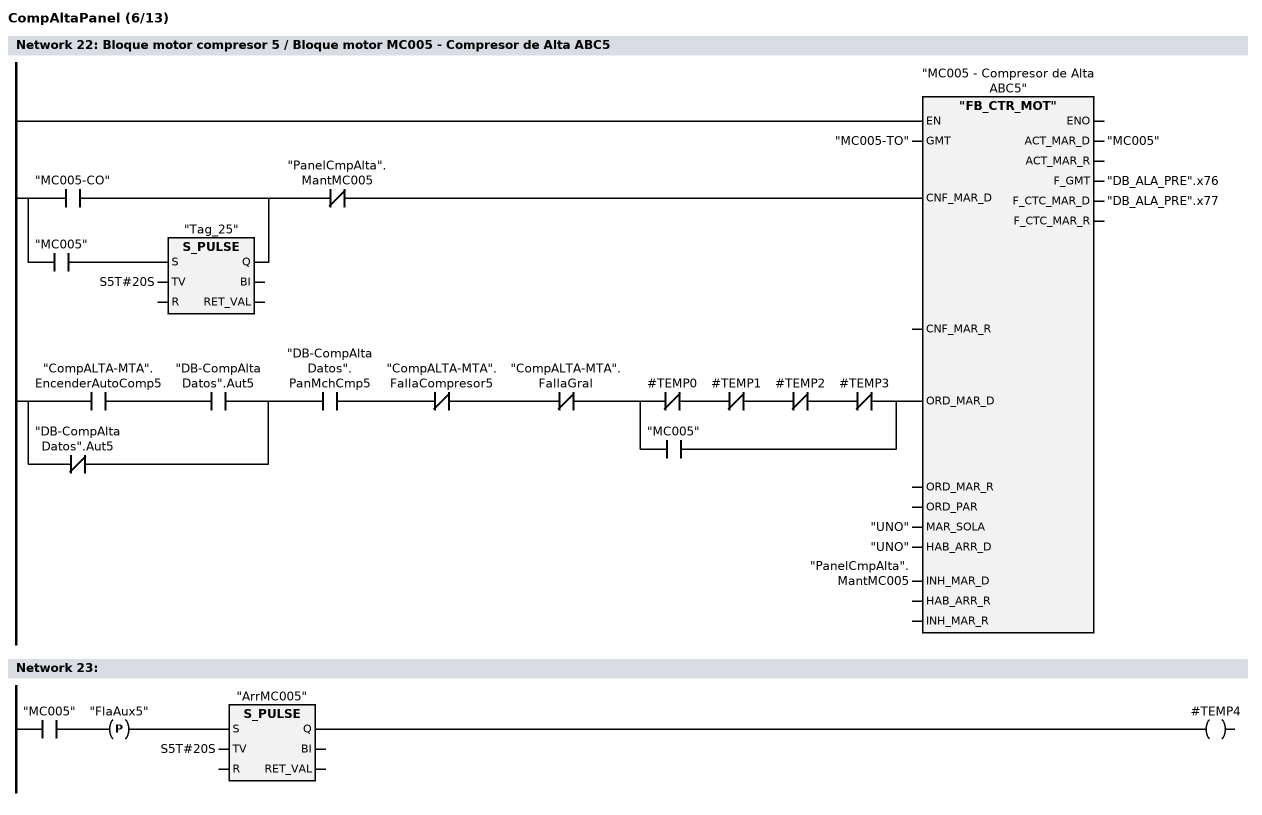
   RUNG wire#powerrail
      "MC005 - Compresor de Alta ABC5"(CNF_MAR_D := wire#w2, ORD_MAR_D := wire#w5, GMT := "MC005-TO", CNF_MAR_R :=, ORD_MAR_R :=, ORD_PAR :=, MAR_SOLA := "UNO", HAB_ARR_D := "UNO", INH_MAR_D := "PanelCmpAlta".MantMC005, HAB_ARR_R :=, INH_MAR_R :=, ACT_MAR_D => "MC005", ACT_MAR_R =>, F_GMT => "DB_ALA_PRE".x76, F_CTC_MAR_D => "DB_ALA_PRE".x77, F_CTC_MAR_R =>)
   END_RUNG
   RUNG wire#powerrail
      Contact( "MC005-CO" )
      wire#w1
      I_Contact( "PanelCmpAlta".MantMC005 )
   END_RUNG wire#w2
   RUNG wire#powerrail
      Contact( "MC005" )
      S_PULSE(T_NO := "Tag_25", TV := S5T#20S, R :=, BI =>, RET_VAL =>)
   END_RUNG wire#w1
   RUNG wire#powerrail
      Contact( "CompALTA-MTA".EncenderAutoComp5 )
      Contact( "DB-CompAltaDatos".Aut5 )
      wire#w3
      Contact( "DB-CompAltaDatos".PanMchCmp5 )
      I_Contact( "CompALTA-MTA".FallaCompresor5 )
      I_Contact( "CompALTA-MTA".FallaGral )
      wire#w4
      I_Contact( #TEMP0 )
      I_Contact( #TEMP1 )
      I_Contact( #TEMP2 )
      I_Contact( #TEMP3 )
   END_RUNG wire#w5
   RUNG wire#powerrail
      I_Contact( "DB-CompAltaDatos".Aut5 )
   END_RUNG wire#w3
   RUNG wire#w4
      Contact( "MC005" )
   END_RUNG wire#w5
   // the same network as SCL:
   #_s5time1 := S_PULSE(T_NO := "Tag_25", S := "MC005", TV := S5T#20S, Q => #_w1);
   "MC005 - Compresor de Alta ABC5"(GMT := "MC005-TO",   // "FB_CTR_MOT"
                           CNF_MAR_D := ("MC005-CO" OR #_w1) AND NOT "PanelCmpAlta".MantMC005,
                           ORD_MAR_D := (("CompALTA-MTA".EncenderAutoComp5 AND "DB-CompAltaDatos".Aut5) OR NOT "DB-CompAltaDatos".Aut5) AND "DB-CompAltaDatos".PanMchCmp5 AND NOT "CompALTA-MTA".FallaCompresor5 AND NOT "CompALTA-MTA".FallaGral AND ((NOT #TEMP0 AND NOT #TEMP1 AND NOT #TEMP2 AND NOT #TEMP3) OR "MC005"),
                           MAR_SOLA := "UNO",
                           HAB_ARR_D := "UNO",
                           INH_MAR_D := "PanelCmpAlta".MantMC005,
                           ACT_MAR_D => "MC005",
                           F_GMT => "DB_ALA_PRE".x76,
                           F_CTC_MAR_D => "DB_ALA_PRE".x77);
END_REGION

REGION Network 23
   RUNG wire#powerrail
      Contact( "MC005" )
      P_Trig( "FlaAux5" )
      S_PULSE(T_NO := "ArrMC005", TV := S5T#20S, R :=, BI =>, RET_VAL =>)
      Coil( #TEMP4 )
   END_RUNG
   // the same network as SCL:
   #_w1 := "MC005" AND NOT "FlaAux5";   // rising edge
   "FlaAux5" := "MC005";
   #_s5time1 := S_PULSE(T_NO := "ArrMC005", S := #_w1, TV := S5T#20S, Q => #_w2);
   #TEMP4 := #_w2;
END_REGION

REGION Network 24: Bloque motor compresor 6 / Bloque motor MC005 - Compresor de Alta ABC5
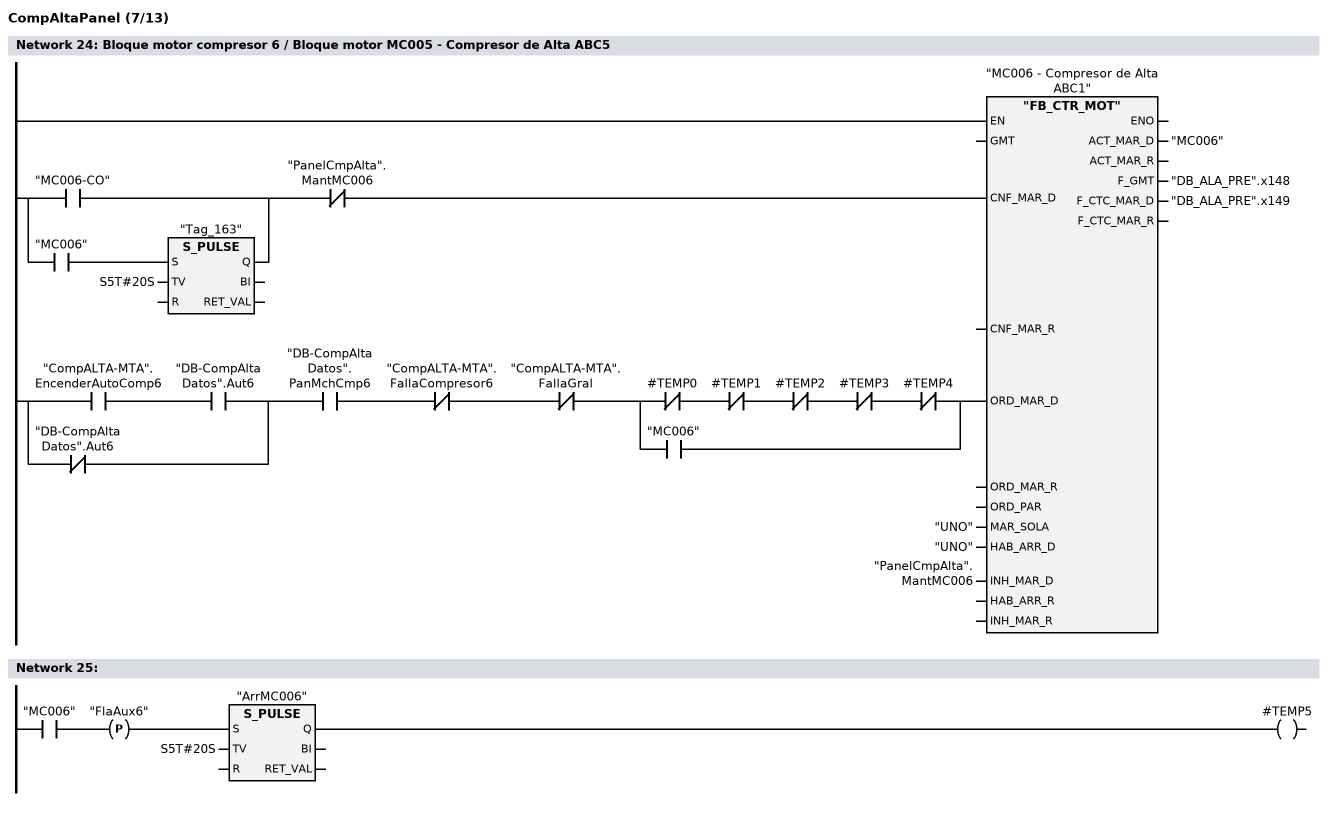
   RUNG wire#powerrail
      "MC006 - Compresor de Alta ABC1"(CNF_MAR_D := wire#w2, ORD_MAR_D := wire#w5, GMT :=, CNF_MAR_R :=, ORD_MAR_R :=, ORD_PAR :=, MAR_SOLA := "UNO", HAB_ARR_D := "UNO", INH_MAR_D := "PanelCmpAlta".MantMC006, HAB_ARR_R :=, INH_MAR_R :=, ACT_MAR_D => "MC006", ACT_MAR_R =>, F_GMT => "DB_ALA_PRE".x148, F_CTC_MAR_D => "DB_ALA_PRE".x149, F_CTC_MAR_R =>)
   END_RUNG
   RUNG wire#powerrail
      Contact( "MC006-CO" )
      wire#w1
      I_Contact( "PanelCmpAlta".MantMC006 )
   END_RUNG wire#w2
   RUNG wire#powerrail
      Contact( "MC006" )
      S_PULSE(T_NO := "Tag_163", TV := S5T#20S, R :=, BI =>, RET_VAL =>)
   END_RUNG wire#w1
   RUNG wire#powerrail
      Contact( "CompALTA-MTA".EncenderAutoComp6 )
      Contact( "DB-CompAltaDatos".Aut6 )
      wire#w3
      Contact( "DB-CompAltaDatos".PanMchCmp6 )
      I_Contact( "CompALTA-MTA".FallaCompresor6 )
      I_Contact( "CompALTA-MTA".FallaGral )
      wire#w4
      I_Contact( #TEMP0 )
      I_Contact( #TEMP1 )
      I_Contact( #TEMP2 )
      I_Contact( #TEMP3 )
      I_Contact( #TEMP4 )
   END_RUNG wire#w5
   RUNG wire#powerrail
      I_Contact( "DB-CompAltaDatos".Aut6 )
   END_RUNG wire#w3
   RUNG wire#w4
      Contact( "MC006" )
   END_RUNG wire#w5
   // the same network as SCL:
   #_s5time1 := S_PULSE(T_NO := "Tag_163", S := "MC006", TV := S5T#20S, Q => #_w1);
   "MC006 - Compresor de Alta ABC1"(CNF_MAR_D := ("MC006-CO" OR #_w1) AND NOT "PanelCmpAlta".MantMC006,   // "FB_CTR_MOT"
                           ORD_MAR_D := (("CompALTA-MTA".EncenderAutoComp6 AND "DB-CompAltaDatos".Aut6) OR NOT "DB-CompAltaDatos".Aut6) AND "DB-CompAltaDatos".PanMchCmp6 AND NOT "CompALTA-MTA".FallaCompresor6 AND NOT "CompALTA-MTA".FallaGral AND ((NOT #TEMP0 AND NOT #TEMP1 AND NOT #TEMP2 AND NOT #TEMP3 AND NOT #TEMP4) OR "MC006"),
                           MAR_SOLA := "UNO",
                           HAB_ARR_D := "UNO",
                           INH_MAR_D := "PanelCmpAlta".MantMC006,
                           ACT_MAR_D => "MC006",
                           F_GMT => "DB_ALA_PRE".x148,
                           F_CTC_MAR_D => "DB_ALA_PRE".x149);
END_REGION

REGION Network 25
   RUNG wire#powerrail
      Contact( "MC006" )
      P_Trig( "FlaAux6" )
      S_PULSE(T_NO := "ArrMC006", TV := S5T#20S, R :=, BI =>, RET_VAL =>)
      Coil( #TEMP5 )
   END_RUNG
   // the same network as SCL:
   #_w1 := "MC006" AND NOT "FlaAux6";   // rising edge
   "FlaAux6" := "MC006";
   #_s5time1 := S_PULSE(T_NO := "ArrMC006", S := #_w1, TV := S5T#20S, Q => #_w2);
   #TEMP5 := #_w2;
END_REGION

REGION Network 26: Bloque de animación motor compresor 1 / Animación Motor MC001 - Compresor de Alta ABC2
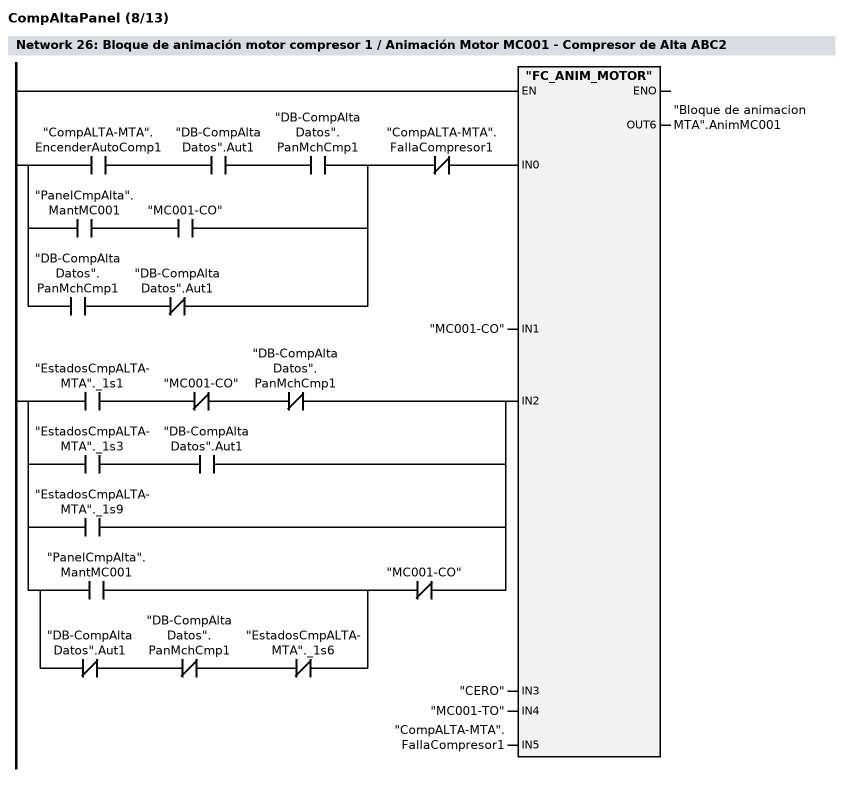
   RUNG wire#powerrail
      "FC_ANIM_MOTOR"(IN0 := wire#w2, IN2 := wire#w4, IN1 := "MC001-CO", IN3 := "CERO", IN4 := "MC001-TO", IN5 := "CompALTA-MTA".FallaCompresor1, OUT6 => "Bloque de animacion MTA".AnimMC001)
   END_RUNG
   RUNG wire#powerrail
      Contact( "CompALTA-MTA".EncenderAutoComp1 )
      Contact( "DB-CompAltaDatos".Aut1 )
      Contact( "DB-CompAltaDatos".PanMchCmp1 )
      wire#w1
      I_Contact( "CompALTA-MTA".FallaCompresor1 )
   END_RUNG wire#w2
   RUNG wire#powerrail
      Contact( "PanelCmpAlta".MantMC001 )
      Contact( "MC001-CO" )
   END_RUNG wire#w1
   RUNG wire#powerrail
      Contact( "DB-CompAltaDatos".PanMchCmp1 )
      I_Contact( "DB-CompAltaDatos".Aut1 )
   END_RUNG wire#w1
   RUNG wire#powerrail
      Contact( "EstadosCmpALTA-MTA"._1s1 )
      I_Contact( "MC001-CO" )
      I_Contact( "DB-CompAltaDatos".PanMchCmp1 )
   END_RUNG wire#w4
   RUNG wire#powerrail
      Contact( "EstadosCmpALTA-MTA"._1s3 )
      Contact( "DB-CompAltaDatos".Aut1 )
   END_RUNG wire#w4
   RUNG wire#powerrail
      Contact( "EstadosCmpALTA-MTA"._1s9 )
   END_RUNG wire#w4
   RUNG wire#powerrail
      Contact( "PanelCmpAlta".MantMC001 )
      wire#w3
      I_Contact( "MC001-CO" )
   END_RUNG wire#w4
   RUNG wire#powerrail
      I_Contact( "DB-CompAltaDatos".Aut1 )
      I_Contact( "DB-CompAltaDatos".PanMchCmp1 )
      I_Contact( "EstadosCmpALTA-MTA"._1s6 )
   END_RUNG wire#w3
   // the same network as SCL:
   "FC_ANIM_MOTOR"(IN0 := (("CompALTA-MTA".EncenderAutoComp1 AND "DB-CompAltaDatos".Aut1 AND "DB-CompAltaDatos".PanMchCmp1) OR ("PanelCmpAlta".MantMC001 AND "MC001-CO") OR ("DB-CompAltaDatos".PanMchCmp1 AND NOT "DB-CompAltaDatos".Aut1)) AND NOT "CompALTA-MTA".FallaCompresor1,
                   IN1 := "MC001-CO",
                   IN2 := ("EstadosCmpALTA-MTA"._1s1 AND NOT "MC001-CO" AND NOT "DB-CompAltaDatos".PanMchCmp1) OR ("EstadosCmpALTA-MTA"._1s3 AND "DB-CompAltaDatos".Aut1) OR "EstadosCmpALTA-MTA"._1s9 OR (("PanelCmpAlta".MantMC001 OR (NOT "DB-CompAltaDatos".Aut1 AND NOT "DB-CompAltaDatos".PanMchCmp1 AND NOT "EstadosCmpALTA-MTA"._1s6)) AND NOT "MC001-CO"),
                   IN3 := "CERO",
                   IN4 := "MC001-TO",
                   IN5 := "CompALTA-MTA".FallaCompresor1,
                   OUT6 => "Bloque de animacion MTA".AnimMC001);
END_REGION

REGION Network 27: Bloque de animación motor compresor 2 / Animación Motor MC002 - Compresor de Alta ABC3
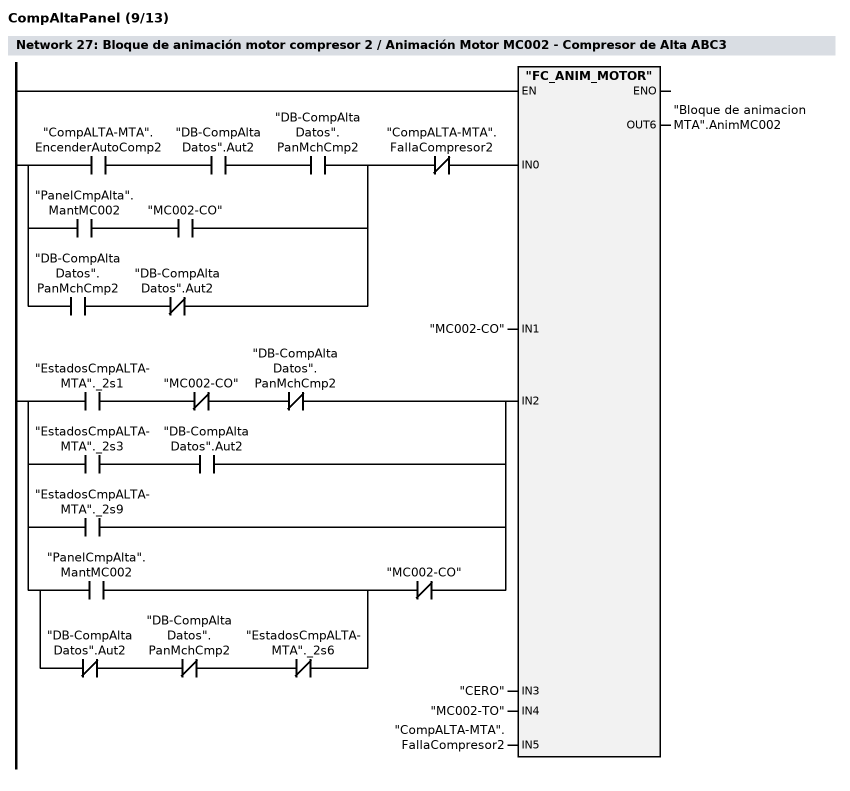
   RUNG wire#powerrail
      "FC_ANIM_MOTOR"(IN0 := wire#w2, IN2 := wire#w4, IN1 := "MC002-CO", IN3 := "CERO", IN4 := "MC002-TO", IN5 := "CompALTA-MTA".FallaCompresor2, OUT6 => "Bloque de animacion MTA".AnimMC002)
   END_RUNG
   RUNG wire#powerrail
      Contact( "CompALTA-MTA".EncenderAutoComp2 )
      Contact( "DB-CompAltaDatos".Aut2 )
      Contact( "DB-CompAltaDatos".PanMchCmp2 )
      wire#w1
      I_Contact( "CompALTA-MTA".FallaCompresor2 )
   END_RUNG wire#w2
   RUNG wire#powerrail
      Contact( "PanelCmpAlta".MantMC002 )
      Contact( "MC002-CO" )
   END_RUNG wire#w1
   RUNG wire#powerrail
      Contact( "DB-CompAltaDatos".PanMchCmp2 )
      I_Contact( "DB-CompAltaDatos".Aut2 )
   END_RUNG wire#w1
   RUNG wire#powerrail
      Contact( "EstadosCmpALTA-MTA"._2s1 )
      I_Contact( "MC002-CO" )
      I_Contact( "DB-CompAltaDatos".PanMchCmp2 )
   END_RUNG wire#w4
   RUNG wire#powerrail
      Contact( "EstadosCmpALTA-MTA"._2s3 )
      Contact( "DB-CompAltaDatos".Aut2 )
   END_RUNG wire#w4
   RUNG wire#powerrail
      Contact( "EstadosCmpALTA-MTA"._2s9 )
   END_RUNG wire#w4
   RUNG wire#powerrail
      Contact( "PanelCmpAlta".MantMC002 )
      wire#w3
      I_Contact( "MC002-CO" )
   END_RUNG wire#w4
   RUNG wire#powerrail
      I_Contact( "DB-CompAltaDatos".Aut2 )
      I_Contact( "DB-CompAltaDatos".PanMchCmp2 )
      I_Contact( "EstadosCmpALTA-MTA"._2s6 )
   END_RUNG wire#w3
   // the same network as SCL:
   "FC_ANIM_MOTOR"(IN0 := (("CompALTA-MTA".EncenderAutoComp2 AND "DB-CompAltaDatos".Aut2 AND "DB-CompAltaDatos".PanMchCmp2) OR ("PanelCmpAlta".MantMC002 AND "MC002-CO") OR ("DB-CompAltaDatos".PanMchCmp2 AND NOT "DB-CompAltaDatos".Aut2)) AND NOT "CompALTA-MTA".FallaCompresor2,
                   IN1 := "MC002-CO",
                   IN2 := ("EstadosCmpALTA-MTA"._2s1 AND NOT "MC002-CO" AND NOT "DB-CompAltaDatos".PanMchCmp2) OR ("EstadosCmpALTA-MTA"._2s3 AND "DB-CompAltaDatos".Aut2) OR "EstadosCmpALTA-MTA"._2s9 OR (("PanelCmpAlta".MantMC002 OR (NOT "DB-CompAltaDatos".Aut2 AND NOT "DB-CompAltaDatos".PanMchCmp2 AND NOT "EstadosCmpALTA-MTA"._2s6)) AND NOT "MC002-CO"),
                   IN3 := "CERO",
                   IN4 := "MC002-TO",
                   IN5 := "CompALTA-MTA".FallaCompresor2,
                   OUT6 => "Bloque de animacion MTA".AnimMC002);
END_REGION

REGION Network 28: Bloque de animación motor compresor 3 / Animación Motor MC003 - Compresor de Alta BELLIS
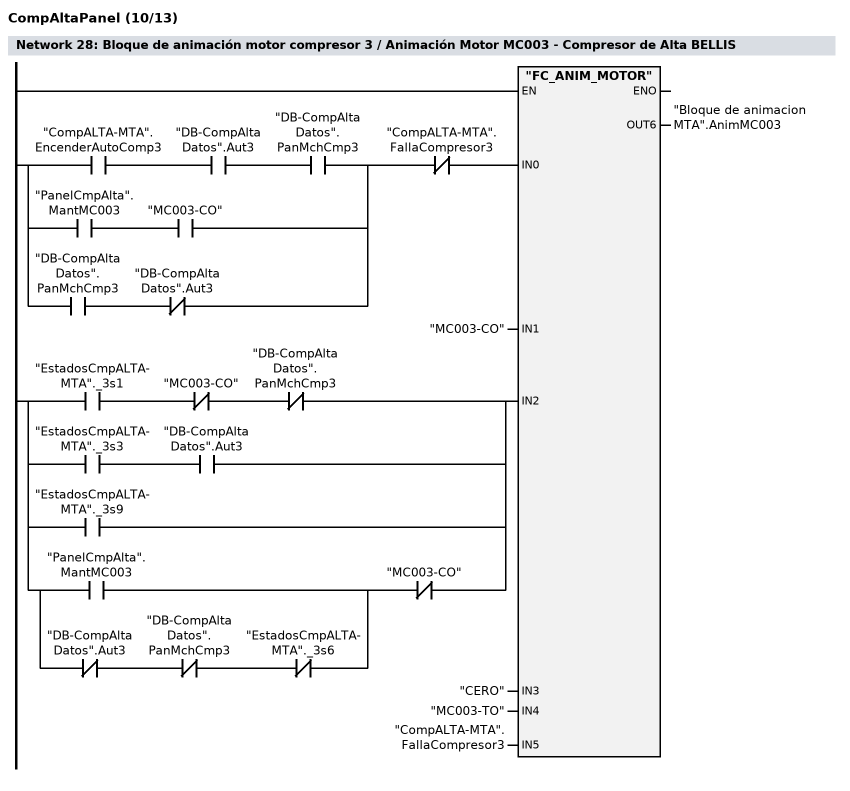
   RUNG wire#powerrail
      "FC_ANIM_MOTOR"(IN0 := wire#w2, IN2 := wire#w4, IN1 := "MC003-CO", IN3 := "CERO", IN4 := "MC003-TO", IN5 := "CompALTA-MTA".FallaCompresor3, OUT6 => "Bloque de animacion MTA".AnimMC003)
   END_RUNG
   RUNG wire#powerrail
      Contact( "CompALTA-MTA".EncenderAutoComp3 )
      Contact( "DB-CompAltaDatos".Aut3 )
      Contact( "DB-CompAltaDatos".PanMchCmp3 )
      wire#w1
      I_Contact( "CompALTA-MTA".FallaCompresor3 )
   END_RUNG wire#w2
   RUNG wire#powerrail
      Contact( "PanelCmpAlta".MantMC003 )
      Contact( "MC003-CO" )
   END_RUNG wire#w1
   RUNG wire#powerrail
      Contact( "DB-CompAltaDatos".PanMchCmp3 )
      I_Contact( "DB-CompAltaDatos".Aut3 )
   END_RUNG wire#w1
   RUNG wire#powerrail
      Contact( "EstadosCmpALTA-MTA"._3s1 )
      I_Contact( "MC003-CO" )
      I_Contact( "DB-CompAltaDatos".PanMchCmp3 )
   END_RUNG wire#w4
   RUNG wire#powerrail
      Contact( "EstadosCmpALTA-MTA"._3s3 )
      Contact( "DB-CompAltaDatos".Aut3 )
   END_RUNG wire#w4
   RUNG wire#powerrail
      Contact( "EstadosCmpALTA-MTA"._3s9 )
   END_RUNG wire#w4
   RUNG wire#powerrail
      Contact( "PanelCmpAlta".MantMC003 )
      wire#w3
      I_Contact( "MC003-CO" )
   END_RUNG wire#w4
   RUNG wire#powerrail
      I_Contact( "DB-CompAltaDatos".Aut3 )
      I_Contact( "DB-CompAltaDatos".PanMchCmp3 )
      I_Contact( "EstadosCmpALTA-MTA"._3s6 )
   END_RUNG wire#w3
   // the same network as SCL:
   "FC_ANIM_MOTOR"(IN0 := (("CompALTA-MTA".EncenderAutoComp3 AND "DB-CompAltaDatos".Aut3 AND "DB-CompAltaDatos".PanMchCmp3) OR ("PanelCmpAlta".MantMC003 AND "MC003-CO") OR ("DB-CompAltaDatos".PanMchCmp3 AND NOT "DB-CompAltaDatos".Aut3)) AND NOT "CompALTA-MTA".FallaCompresor3,
                   IN1 := "MC003-CO",
                   IN2 := ("EstadosCmpALTA-MTA"._3s1 AND NOT "MC003-CO" AND NOT "DB-CompAltaDatos".PanMchCmp3) OR ("EstadosCmpALTA-MTA"._3s3 AND "DB-CompAltaDatos".Aut3) OR "EstadosCmpALTA-MTA"._3s9 OR (("PanelCmpAlta".MantMC003 OR (NOT "DB-CompAltaDatos".Aut3 AND NOT "DB-CompAltaDatos".PanMchCmp3 AND NOT "EstadosCmpALTA-MTA"._3s6)) AND NOT "MC003-CO"),
                   IN3 := "CERO",
                   IN4 := "MC003-TO",
                   IN5 := "CompALTA-MTA".FallaCompresor3,
                   OUT6 => "Bloque de animacion MTA".AnimMC003);
END_REGION

REGION Network 29: Bloque de animación motor compresor 4 / Animación Motor MC004 - Compresor de Alta ABC4
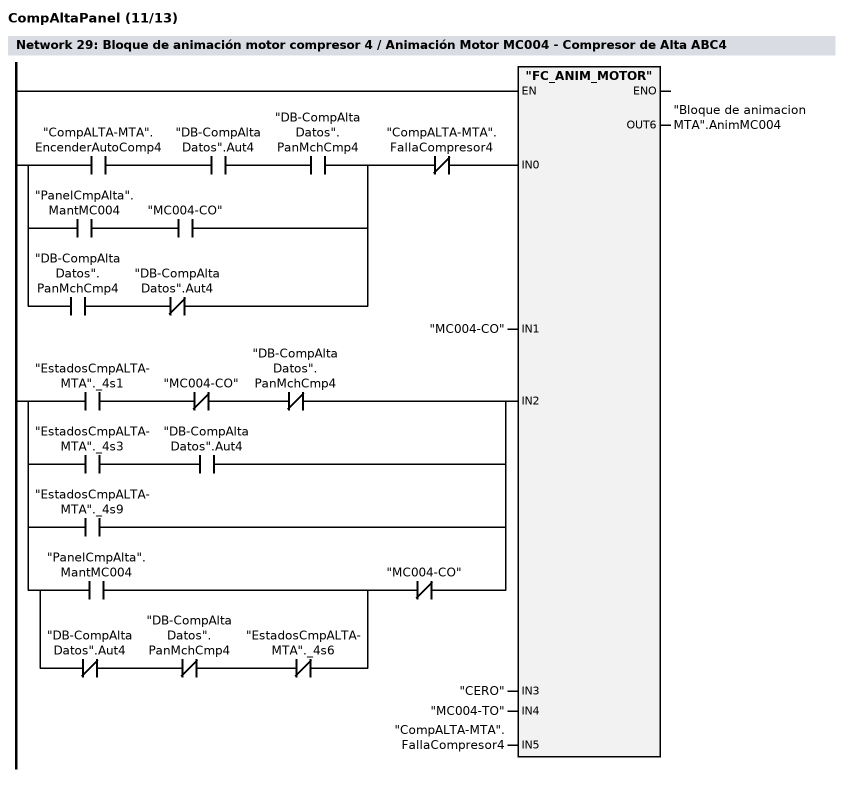
   RUNG wire#powerrail
      "FC_ANIM_MOTOR"(IN0 := wire#w2, IN2 := wire#w4, IN1 := "MC004-CO", IN3 := "CERO", IN4 := "MC004-TO", IN5 := "CompALTA-MTA".FallaCompresor4, OUT6 => "Bloque de animacion MTA".AnimMC004)
   END_RUNG
   RUNG wire#powerrail
      Contact( "CompALTA-MTA".EncenderAutoComp4 )
      Contact( "DB-CompAltaDatos".Aut4 )
      Contact( "DB-CompAltaDatos".PanMchCmp4 )
      wire#w1
      I_Contact( "CompALTA-MTA".FallaCompresor4 )
   END_RUNG wire#w2
   RUNG wire#powerrail
      Contact( "PanelCmpAlta".MantMC004 )
      Contact( "MC004-CO" )
   END_RUNG wire#w1
   RUNG wire#powerrail
      Contact( "DB-CompAltaDatos".PanMchCmp4 )
      I_Contact( "DB-CompAltaDatos".Aut4 )
   END_RUNG wire#w1
   RUNG wire#powerrail
      Contact( "EstadosCmpALTA-MTA"._4s1 )
      I_Contact( "MC004-CO" )
      I_Contact( "DB-CompAltaDatos".PanMchCmp4 )
   END_RUNG wire#w4
   RUNG wire#powerrail
      Contact( "EstadosCmpALTA-MTA"._4s3 )
      Contact( "DB-CompAltaDatos".Aut4 )
   END_RUNG wire#w4
   RUNG wire#powerrail
      Contact( "EstadosCmpALTA-MTA"._4s9 )
   END_RUNG wire#w4
   RUNG wire#powerrail
      Contact( "PanelCmpAlta".MantMC004 )
      wire#w3
      I_Contact( "MC004-CO" )
   END_RUNG wire#w4
   RUNG wire#powerrail
      I_Contact( "DB-CompAltaDatos".Aut4 )
      I_Contact( "DB-CompAltaDatos".PanMchCmp4 )
      I_Contact( "EstadosCmpALTA-MTA"._4s6 )
   END_RUNG wire#w3
   // the same network as SCL:
   "FC_ANIM_MOTOR"(IN0 := (("CompALTA-MTA".EncenderAutoComp4 AND "DB-CompAltaDatos".Aut4 AND "DB-CompAltaDatos".PanMchCmp4) OR ("PanelCmpAlta".MantMC004 AND "MC004-CO") OR ("DB-CompAltaDatos".PanMchCmp4 AND NOT "DB-CompAltaDatos".Aut4)) AND NOT "CompALTA-MTA".FallaCompresor4,
                   IN1 := "MC004-CO",
                   IN2 := ("EstadosCmpALTA-MTA"._4s1 AND NOT "MC004-CO" AND NOT "DB-CompAltaDatos".PanMchCmp4) OR ("EstadosCmpALTA-MTA"._4s3 AND "DB-CompAltaDatos".Aut4) OR "EstadosCmpALTA-MTA"._4s9 OR (("PanelCmpAlta".MantMC004 OR (NOT "DB-CompAltaDatos".Aut4 AND NOT "DB-CompAltaDatos".PanMchCmp4 AND NOT "EstadosCmpALTA-MTA"._4s6)) AND NOT "MC004-CO"),
                   IN3 := "CERO",
                   IN4 := "MC004-TO",
                   IN5 := "CompALTA-MTA".FallaCompresor4,
                   OUT6 => "Bloque de animacion MTA".AnimMC004);
END_REGION

REGION Network 30: Bloque de animación motor compresor 5 / Animación Motor MC005 - Compresor de Alta ABC5
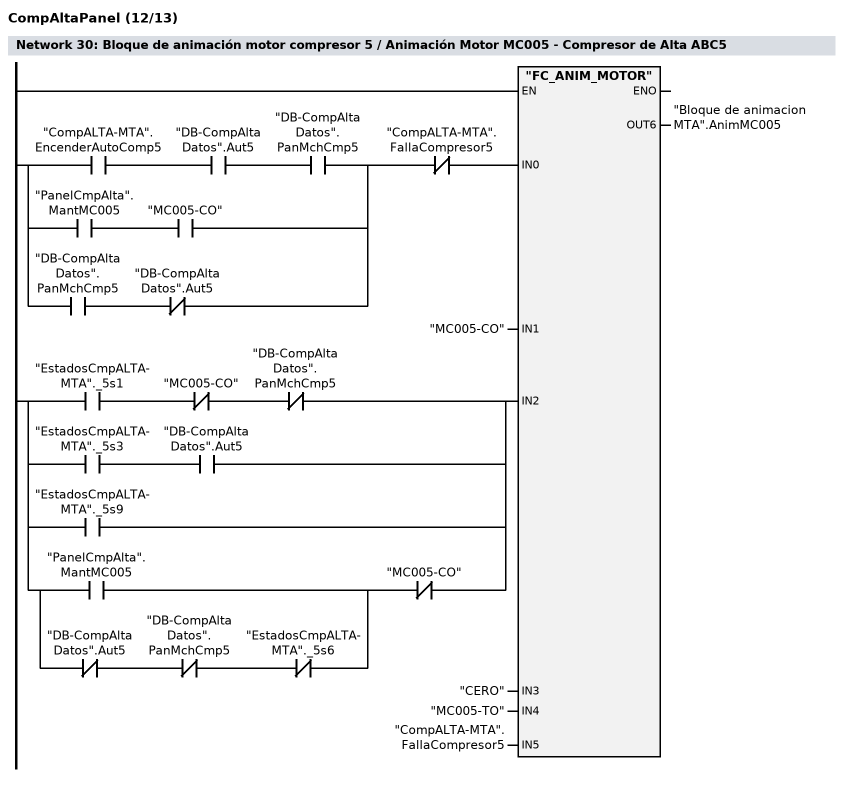
   RUNG wire#powerrail
      "FC_ANIM_MOTOR"(IN0 := wire#w2, IN2 := wire#w4, IN1 := "MC005-CO", IN3 := "CERO", IN4 := "MC005-TO", IN5 := "CompALTA-MTA".FallaCompresor5, OUT6 => "Bloque de animacion MTA".AnimMC005)
   END_RUNG
   RUNG wire#powerrail
      Contact( "CompALTA-MTA".EncenderAutoComp5 )
      Contact( "DB-CompAltaDatos".Aut5 )
      Contact( "DB-CompAltaDatos".PanMchCmp5 )
      wire#w1
      I_Contact( "CompALTA-MTA".FallaCompresor5 )
   END_RUNG wire#w2
   RUNG wire#powerrail
      Contact( "PanelCmpAlta".MantMC005 )
      Contact( "MC005-CO" )
   END_RUNG wire#w1
   RUNG wire#powerrail
      Contact( "DB-CompAltaDatos".PanMchCmp5 )
      I_Contact( "DB-CompAltaDatos".Aut5 )
   END_RUNG wire#w1
   RUNG wire#powerrail
      Contact( "EstadosCmpALTA-MTA"._5s1 )
      I_Contact( "MC005-CO" )
      I_Contact( "DB-CompAltaDatos".PanMchCmp5 )
   END_RUNG wire#w4
   RUNG wire#powerrail
      Contact( "EstadosCmpALTA-MTA"._5s3 )
      Contact( "DB-CompAltaDatos".Aut5 )
   END_RUNG wire#w4
   RUNG wire#powerrail
      Contact( "EstadosCmpALTA-MTA"._5s9 )
   END_RUNG wire#w4
   RUNG wire#powerrail
      Contact( "PanelCmpAlta".MantMC005 )
      wire#w3
      I_Contact( "MC005-CO" )
   END_RUNG wire#w4
   RUNG wire#powerrail
      I_Contact( "DB-CompAltaDatos".Aut5 )
      I_Contact( "DB-CompAltaDatos".PanMchCmp5 )
      I_Contact( "EstadosCmpALTA-MTA"._5s6 )
   END_RUNG wire#w3
   // the same network as SCL:
   "FC_ANIM_MOTOR"(IN0 := (("CompALTA-MTA".EncenderAutoComp5 AND "DB-CompAltaDatos".Aut5 AND "DB-CompAltaDatos".PanMchCmp5) OR ("PanelCmpAlta".MantMC005 AND "MC005-CO") OR ("DB-CompAltaDatos".PanMchCmp5 AND NOT "DB-CompAltaDatos".Aut5)) AND NOT "CompALTA-MTA".FallaCompresor5,
                   IN1 := "MC005-CO",
                   IN2 := ("EstadosCmpALTA-MTA"._5s1 AND NOT "MC005-CO" AND NOT "DB-CompAltaDatos".PanMchCmp5) OR ("EstadosCmpALTA-MTA"._5s3 AND "DB-CompAltaDatos".Aut5) OR "EstadosCmpALTA-MTA"._5s9 OR (("PanelCmpAlta".MantMC005 OR (NOT "DB-CompAltaDatos".Aut5 AND NOT "DB-CompAltaDatos".PanMchCmp5 AND NOT "EstadosCmpALTA-MTA"._5s6)) AND NOT "MC005-CO"),
                   IN3 := "CERO",
                   IN4 := "MC005-TO",
                   IN5 := "CompALTA-MTA".FallaCompresor5,
                   OUT6 => "Bloque de animacion MTA".AnimMC005);
END_REGION

REGION Network 31: Bloque de animación motor compresor 6 / Animación Motor MC005 - Compresor de Alta ABC5
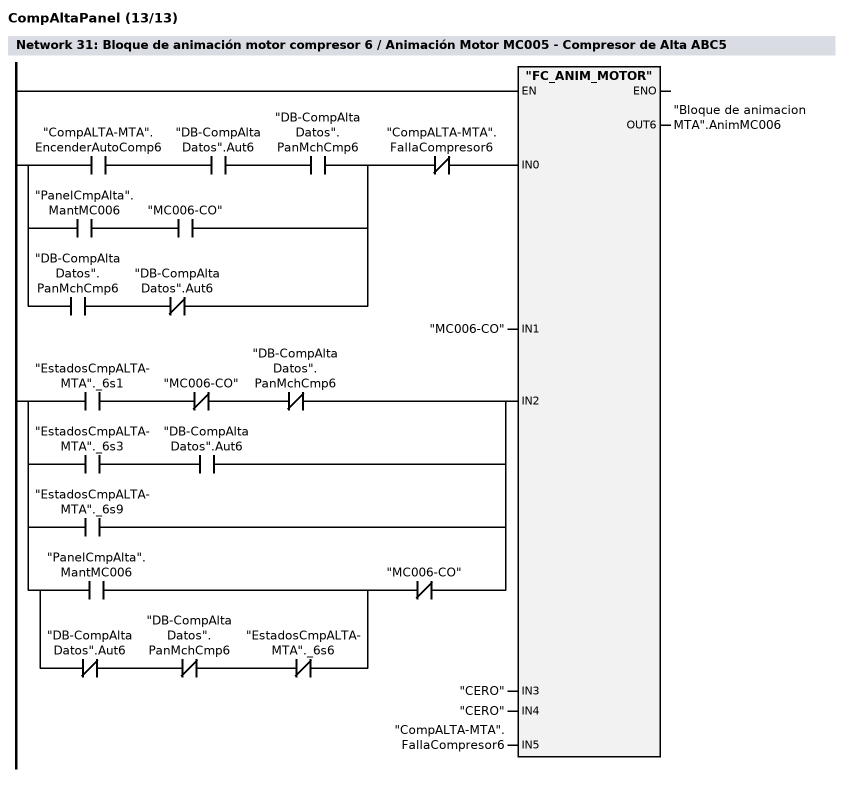
   RUNG wire#powerrail
      "FC_ANIM_MOTOR"(IN0 := wire#w2, IN2 := wire#w4, IN1 := "MC006-CO", IN3 := "CERO", IN4 := "CERO", IN5 := "CompALTA-MTA".FallaCompresor6, OUT6 => "Bloque de animacion MTA".AnimMC006)
   END_RUNG
   RUNG wire#powerrail
      Contact( "CompALTA-MTA".EncenderAutoComp6 )
      Contact( "DB-CompAltaDatos".Aut6 )
      Contact( "DB-CompAltaDatos".PanMchCmp6 )
      wire#w1
      I_Contact( "CompALTA-MTA".FallaCompresor6 )
   END_RUNG wire#w2
   RUNG wire#powerrail
      Contact( "PanelCmpAlta".MantMC006 )
      Contact( "MC006-CO" )
   END_RUNG wire#w1
   RUNG wire#powerrail
      Contact( "DB-CompAltaDatos".PanMchCmp6 )
      I_Contact( "DB-CompAltaDatos".Aut6 )
   END_RUNG wire#w1
   RUNG wire#powerrail
      Contact( "EstadosCmpALTA-MTA"._6s1 )
      I_Contact( "MC006-CO" )
      I_Contact( "DB-CompAltaDatos".PanMchCmp6 )
   END_RUNG wire#w4
   RUNG wire#powerrail
      Contact( "EstadosCmpALTA-MTA"._6s3 )
      Contact( "DB-CompAltaDatos".Aut6 )
   END_RUNG wire#w4
   RUNG wire#powerrail
      Contact( "EstadosCmpALTA-MTA"._6s9 )
   END_RUNG wire#w4
   RUNG wire#powerrail
      Contact( "PanelCmpAlta".MantMC006 )
      wire#w3
      I_Contact( "MC006-CO" )
   END_RUNG wire#w4
   RUNG wire#powerrail
      I_Contact( "DB-CompAltaDatos".Aut6 )
      I_Contact( "DB-CompAltaDatos".PanMchCmp6 )
      I_Contact( "EstadosCmpALTA-MTA"._6s6 )
   END_RUNG wire#w3
   // the same network as SCL:
   "FC_ANIM_MOTOR"(IN0 := (("CompALTA-MTA".EncenderAutoComp6 AND "DB-CompAltaDatos".Aut6 AND "DB-CompAltaDatos".PanMchCmp6) OR ("PanelCmpAlta".MantMC006 AND "MC006-CO") OR ("DB-CompAltaDatos".PanMchCmp6 AND NOT "DB-CompAltaDatos".Aut6)) AND NOT "CompALTA-MTA".FallaCompresor6,
                   IN1 := "MC006-CO",
                   IN2 := ("EstadosCmpALTA-MTA"._6s1 AND NOT "MC006-CO" AND NOT "DB-CompAltaDatos".PanMchCmp6) OR ("EstadosCmpALTA-MTA"._6s3 AND "DB-CompAltaDatos".Aut6) OR "EstadosCmpALTA-MTA"._6s9 OR (("PanelCmpAlta".MantMC006 OR (NOT "DB-CompAltaDatos".Aut6 AND NOT "DB-CompAltaDatos".PanMchCmp6 AND NOT "EstadosCmpALTA-MTA"._6s6)) AND NOT "MC006-CO"),
                   IN3 := "CERO",
                   IN4 := "CERO",
                   IN5 := "CompALTA-MTA".FallaCompresor6,
                   OUT6 => "Bloque de animacion MTA".AnimMC006);
END_REGION
END_FUNCTION

FUNCTION "ModoManualAlta" : Void   // FC48, LAD
{ S7_Optimized_Access := 'FALSE' }
VERSION : 0.1
   VAR_TEMP   // added for the SCL form of the ladder/FBD networks
      _w1 : Bool;
      _s5time1 : S5Time;
   END_VAR
BEGIN

REGION Network 1
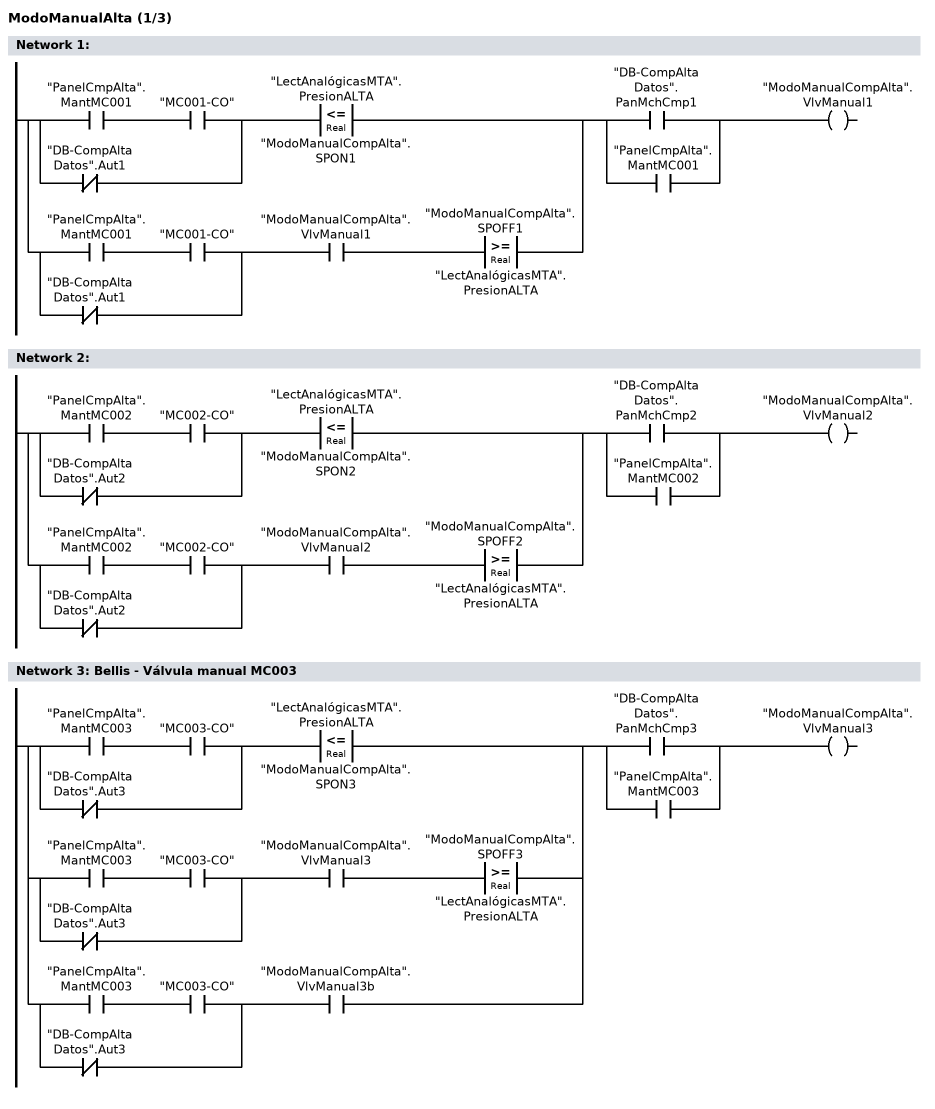
   "ModoManualCompAlta".VlvManual1 := (((NOT "DB-CompAltaDatos".Aut1 OR ("PanelCmpAlta".MantMC001 AND "MC001-CO")) AND ("LectAnalógicasMTA".PresionALTA <= "ModoManualCompAlta".SPON1)) OR ((NOT "DB-CompAltaDatos".Aut1 OR ("PanelCmpAlta".MantMC001 AND "MC001-CO")) AND "ModoManualCompAlta".VlvManual1 AND ("ModoManualCompAlta".SPOFF1 >= "LectAnalógicasMTA".PresionALTA))) AND ("DB-CompAltaDatos".PanMchCmp1 OR "PanelCmpAlta".MantMC001);
END_REGION

REGION Network 2
   "ModoManualCompAlta".VlvManual2 := (((NOT "DB-CompAltaDatos".Aut2 OR ("PanelCmpAlta".MantMC002 AND "MC002-CO")) AND ("LectAnalógicasMTA".PresionALTA <= "ModoManualCompAlta".SPON2)) OR ((NOT "DB-CompAltaDatos".Aut2 OR ("PanelCmpAlta".MantMC002 AND "MC002-CO")) AND "ModoManualCompAlta".VlvManual2 AND ("ModoManualCompAlta".SPOFF2 >= "LectAnalógicasMTA".PresionALTA))) AND ("DB-CompAltaDatos".PanMchCmp2 OR "PanelCmpAlta".MantMC002);
END_REGION

REGION Network 3: Bellis - Válvula manual MC003
   "ModoManualCompAlta".VlvManual3 := (((NOT "DB-CompAltaDatos".Aut3 OR ("PanelCmpAlta".MantMC003 AND "MC003-CO")) AND ("LectAnalógicasMTA".PresionALTA <= "ModoManualCompAlta".SPON3)) OR ((NOT "DB-CompAltaDatos".Aut3 OR ("PanelCmpAlta".MantMC003 AND "MC003-CO")) AND "ModoManualCompAlta".VlvManual3 AND ("ModoManualCompAlta".SPOFF3 >= "LectAnalógicasMTA".PresionALTA)) OR ((NOT "DB-CompAltaDatos".Aut3 OR ("PanelCmpAlta".MantMC003 AND "MC003-CO")) AND "ModoManualCompAlta".VlvManual3b)) AND ("DB-CompAltaDatos".PanMchCmp3 OR "PanelCmpAlta".MantMC003);
END_REGION

REGION Network 4: Bellis - Válvula manual MC003b